// TIA Portal project "PolyMix_v0.1" (V14) (continued)
VERSION : 0.1
   VAR
      DD_Status : Int;
      DD_Mode : Int;
      DD_Alarm : Word;
      DL_Status : Int;
      DL_Mode : Int;
      DL_Alarm : Word;
      Mix_1_Status : Int;
      Mix_1_Mode : Int;
      Mix_1_Alarm : Word;
      Mix_2_Status : Int;
      Mix_2_Mode : Int;
      Mix_2_Alarm : Word;
      Mix_3_Status : Int;
      Mix_3_Mode : Int;
      Mix_3_Alarm : Word;
      KC1_Status : Int;
      Flowmeter : Real;
      Flow_Alarm : Word;
      Level : Real;
      Level_Alarm : Word;
      SP : Real;
      Start : Bool;
      Hand : Bool;
      Warning : Bool;
      Config : Struct
         Use_DD : Bool;   // Использовать сухой дозатор
         Use_DL : Bool;   // Использовать жидкий дозатор
         Use_Mix_1 : Bool;   // Использовать мешалку 1
         Use_Mix_2 : Bool;   // Использовать мешалку 2
         Use_Mix_3 : Bool;   // Использовать мешалку 3
      END_STRUCT;
      Alarm : Word;
   END_VAR
BEGIN
END_DATA_BLOCK

DATA_BLOCK "Time"   // DB13
{ S7_Optimized_Access := 'FALSE' }
VERSION : 0.1
   VAR
      Today : DTL;
      Today_status : Int;
      Set_DTL : DTL;
      Set_status : Int;
      Year : UInt;
      Month : UInt;
      Day : UInt;
      Hour : UInt;
      Minutes : UInt;
      Save : Bool;   // Сохранить время
   END_VAR
BEGIN
END_DATA_BLOCK

// folder: Modules

DATA_BLOCK "DIx_DB"   // DB200
{ S7_Optimized_Access := 'FALSE' }
VERSION : 0.1
// stored: InstanceOfName DIx
"DIx"
BEGIN
END_DATA_BLOCK

DATA_BLOCK "DOx_DB"   // DB201
{ S7_Optimized_Access := 'FALSE' }
VERSION : 0.1
// stored: InstanceOfName DOx
"DOx"
BEGIN
END_DATA_BLOCK

// folder: System blocks/Program resources

DATA_BLOCK "T_Reset"   // DB7
{ S7_Optimized_Access := 'TRUE' }
AUTHOR : Simatic
FAMILY : IEC
NAME : IEC_TMR
VERSION : 1.0
// stored: InstanceOfName IEC_TIMER
"IEC_TIMER"
BEGIN
END_DATA_BLOCK

DATA_BLOCK "clock_5s_ON"   // DB507
{ S7_Optimized_Access := 'TRUE' }
AUTHOR : Simatic
FAMILY : IEC
NAME : IEC_TMR
VERSION : 1.0
// stored: InstanceOfName IEC_TIMER
"IEC_TIMER"
BEGIN
END_DATA_BLOCK

DATA_BLOCK "clock_5s_OFF"   // DB508
{ S7_Optimized_Access := 'TRUE' }
AUTHOR : Simatic
FAMILY : IEC
NAME : IEC_TMR
VERSION : 1.0
// stored: InstanceOfName IEC_TIMER
"IEC_TIMER"
BEGIN
END_DATA_BLOCK

// folder: (top level)

ORGANIZATION_BLOCK "Main"   // OB1, LAD, ProgramCycle
TITLE = "Main Program Sweep (Cycle)"
{ S7_Optimized_Access := 'TRUE' }
VERSION : 0.1
   VAR_INPUT
      Initial_Call : Bool;   // Initial call of this OB
      Remanence : Bool;   // =True, if remanent data are available
   END_VAR
   VAR_TEMP   // added for the SCL form of the ladder/FBD networks
      _w1 : Bool;
   END_VAR
BEGIN

REGION Network 1
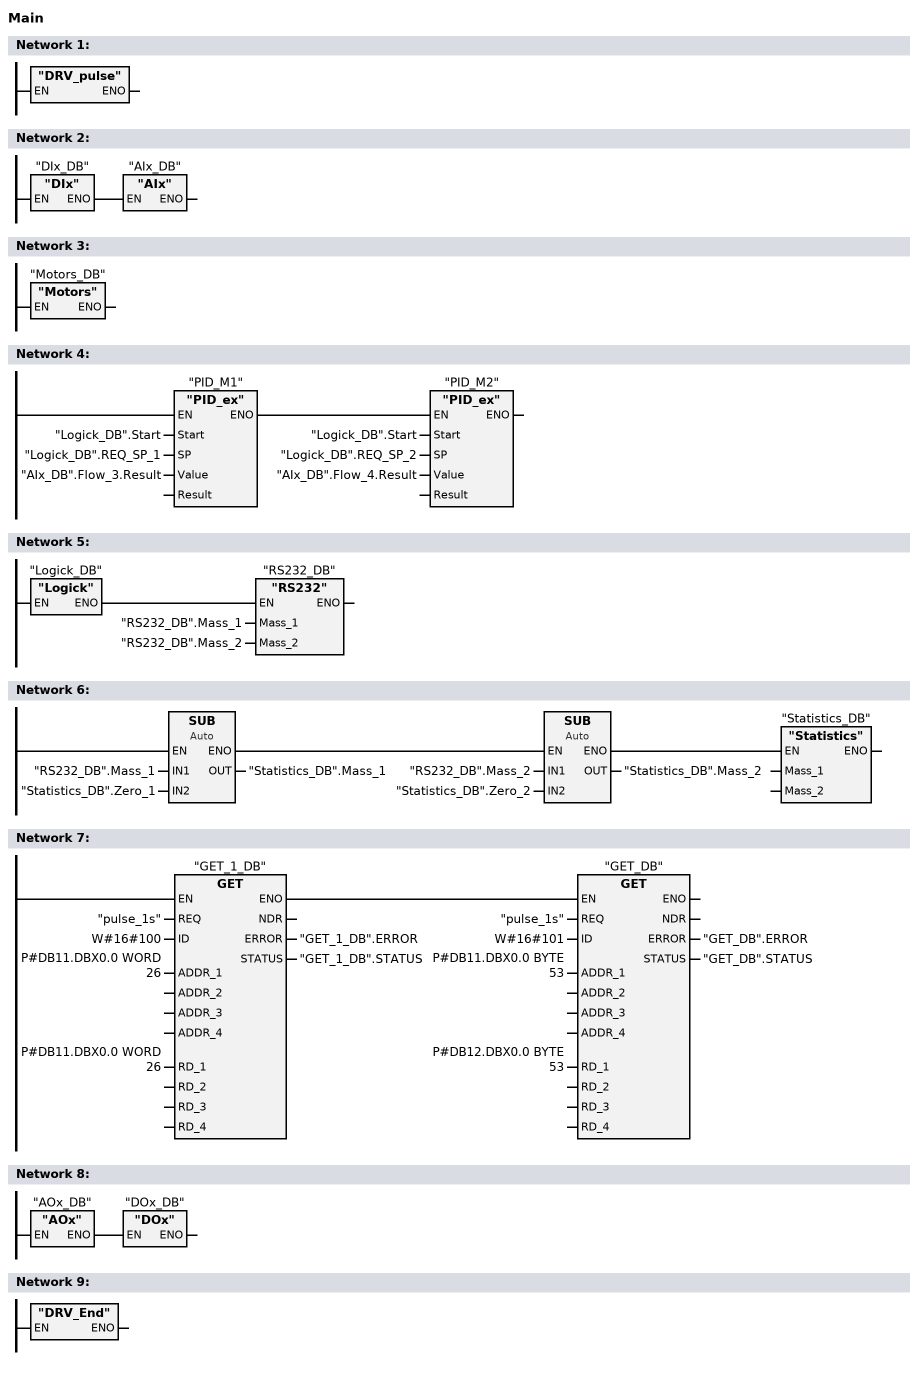
   RUNG wire#powerrail
      "DRV_pulse"()
   END_RUNG
   // the same network as SCL:
   "DRV_pulse"();
END_REGION

REGION Network 2
   RUNG wire#powerrail
      "DIx_DB"()
      "AIx_DB"()
   END_RUNG
   // the same network as SCL:
   "DIx_DB"(ENO => #_w1);   // "DIx"
   IF #_w1 THEN
       "AIx_DB"();   // "AIx"
   END_IF;
END_REGION

REGION Network 3
   RUNG wire#powerrail
      "Motors_DB"()
   END_RUNG
   // the same network as SCL:
   "Motors_DB"();   // "Motors"
END_REGION

REGION Network 4
   RUNG wire#powerrail
      "PID_M1"(Start := "Logick_DB".Start, SP := "Logick_DB".REQ_SP_1, Value := "AIx_DB".Flow_3.Result, Result :=)
      "PID_M2"(Start := "Logick_DB".Start, SP := "Logick_DB".REQ_SP_2, Value := "AIx_DB".Flow_4.Result, Result :=)
   END_RUNG
   // the same network as SCL:
   "PID_M1"(Start := "Logick_DB".Start,   // "PID_ex"
            SP := "Logick_DB".REQ_SP_1,
            Value := "AIx_DB".Flow_3.Result,
            ENO => #_w1);
   IF #_w1 THEN
       "PID_M2"(Start := "Logick_DB".Start, SP := "Logick_DB".REQ_SP_2, Value := "AIx_DB".Flow_4.Result);   // "PID_ex"
   END_IF;
END_REGION

REGION Network 5
   RUNG wire#powerrail
      "Logick_DB"()
      "RS232_DB"(Mass_1 := "RS232_DB".Mass_1, Mass_2 := "RS232_DB".Mass_2)
   END_RUNG
   // the same network as SCL:
   "Logick_DB"(ENO => #_w1);   // "Logick"
   IF #_w1 THEN
       "RS232_DB"(Mass_1 := "RS232_DB".Mass_1, Mass_2 := "RS232_DB".Mass_2);   // "RS232"
   END_IF;
END_REGION

REGION Network 6
   RUNG wire#powerrail
      Sub(in1 := "RS232_DB".Mass_1, in2 := "Statistics_DB".Zero_1, out => "Statistics_DB".Mass_1)
      Sub(in1 := "RS232_DB".Mass_2, in2 := "Statistics_DB".Zero_2, out => "Statistics_DB".Mass_2)
      "Statistics_DB"(Mass_1 :=, Mass_2 :=)
   END_RUNG
   // the same network as SCL:
   "Statistics_DB".Mass_1 := "RS232_DB".Mass_1 - "Statistics_DB".Zero_1;
   "Statistics_DB".Mass_2 := "RS232_DB".Mass_2 - "Statistics_DB".Zero_2;
   "Statistics_DB"();   // "Statistics"
END_REGION

REGION Network 7
   // ENO of a box is taken as its EN; it also drops when the box reports an error
   "GET_1_DB"(REQ := "pulse_1s",   // GET
              ID := W#16#100,
              ADDR_1 := P#DB11.DBX0.0 WORD 26,
              RD_1 := P#DB11.DBX0.0 WORD 26,
              ERROR => "GET_1_DB".ERROR,
              STATUS => "GET_1_DB".STATUS);
   "GET_DB"(REQ := "pulse_1s",   // GET
            ID := W#16#101,
            ADDR_1 := P#DB11.DBX0.0 BYTE 53,
            RD_1 := P#DB12.DBX0.0 BYTE 53,
            ERROR => "GET_DB".ERROR,
            STATUS => "GET_DB".STATUS);
END_REGION

REGION Network 8
   RUNG wire#powerrail
      "AOx_DB"()
      "DOx_DB"()
   END_RUNG
   // the same network as SCL:
   "AOx_DB"(ENO => #_w1);   // "AOx"
   IF #_w1 THEN
       "DOx_DB"();   // "DOx"
   END_IF;
END_REGION

REGION Network 9
   RUNG wire#powerrail
      "DRV_End"()
   END_RUNG
   // the same network as SCL:
   "DRV_End"();
END_REGION
END_ORGANIZATION_BLOCK

ORGANIZATION_BLOCK "Time error interrupt"   // OB80, LAD, TimeErrorInterrupt
{ S7_Optimized_Access := 'TRUE' }
VERSION : 0.1
   VAR_INPUT
      Fault_ID : Byte;   // Fault identifier
      Csg_OBnr : OB_Any;   // Number of OB causing the error
      Csg_Prio : UInt;   // Priority of OB causing the error
   END_VAR
BEGIN
END_ORGANIZATION_BLOCK

ORGANIZATION_BLOCK "Diagnostic error interrupt"   // OB82, LAD, DiagnosticErrorInterrupt
{ S7_Optimized_Access := 'TRUE' }
VERSION : 0.1
   VAR_INPUT
      IO_State : Word;   // IO state of the HW object
      LADDR : Hw_Any;   // Hardware identifier
      Channel : UInt;   // Channel number
      MultiError : Bool;   // =true if more than one error is present
   END_VAR
BEGIN
END_ORGANIZATION_BLOCK

ORGANIZATION_BLOCK "Startup"   // OB100, LAD, Startup
TITLE = "Complete Restart"
{ S7_Optimized_Access := 'TRUE' }
VERSION : 0.1
   VAR_INPUT
      LostRetentive : Bool;   // True if retentive data are lost
      LostRTC : Bool;   // True if date and time are lost
   END_VAR
BEGIN

REGION Network 1: Запуск автоматики
END_REGION

REGION Network 2
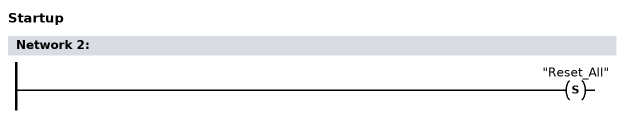
   RUNG wire#powerrail
      S_Coil( "Reset_All" )
   END_RUNG
   // the same network as SCL:
   "Reset_All" := TRUE;
END_REGION
END_ORGANIZATION_BLOCK

// folder: DRV_Low

FUNCTION_BLOCK "DI_ex"   // FB100, LAD
{ S7_Optimized_Access := 'FALSE' }
VERSION : 0.1
   VAR_INPUT
      Input : Bool;   // Входящий сигнал
      pulse : Bool;   // Частота фильтрации дребезка
   END_VAR
   VAR_OUTPUT
      Signal : Bool;   // Результирующий сигнал
   END_VAR
   VAR
      Hand : Bool;   // 0 - Авто, 1 - Ручной
      Start_M : Bool;   // Запуск в ручном режиме
      Data : Bool;   // Отфильтрованный сигнал
      Inverse : Bool;   // Инверсия входного сигнала
      Filter_On : Struct   // Фильтр наличия сигнала
         SP : Int;
         Now : Int;
         "Exit" : Bool;
         Start : Bool;
         Pause : Bool;
         Reset : Bool;
      END_STRUCT;
      Filter_Off : Struct   // Фильтр отсутствия сигнала
         SP : Int;
         Now : Int;
         "Exit" : Bool;
         Start : Bool;
         Pause : Bool;
         Reset : Bool;
      END_STRUCT;
      res_1 : Word;
   END_VAR
   VAR_TEMP   // added for the SCL form of the ladder/FBD networks
      _w1 : Bool;
   END_VAR
BEGIN

REGION Network 1: Устройство в ручном режиме
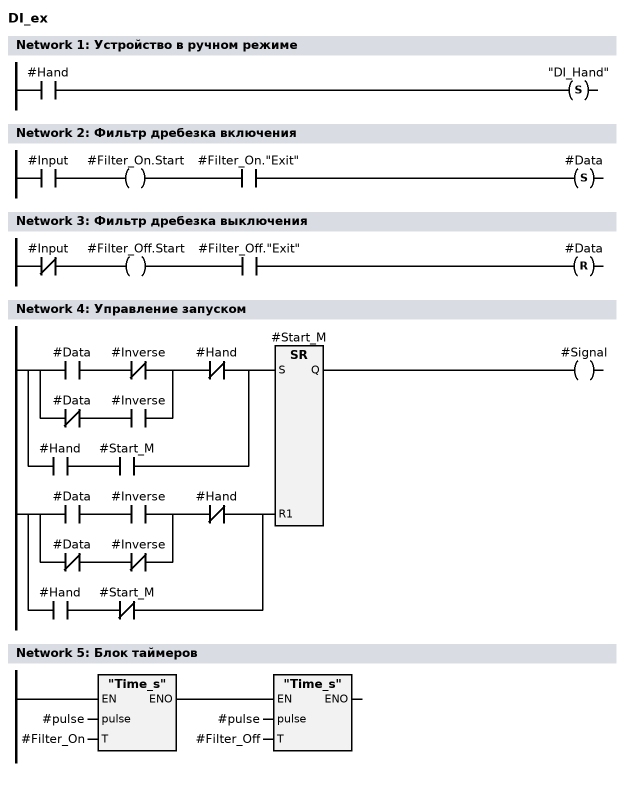
   RUNG wire#powerrail
      Contact( #Hand )
      S_Coil( "DI_Hand" )
   END_RUNG
   // the same network as SCL:
   IF #Hand THEN "DI_Hand" := TRUE; END_IF;
END_REGION

REGION Network 2: Фильтр дребезка включения
   RUNG wire#powerrail
      Contact( #Input )
      Coil( #Filter_On.Start )
      Contact( #Filter_On."Exit" )
      S_Coil( #Data )
   END_RUNG
   // the same network as SCL:
   #Filter_On.Start := #Input;
   IF #Input AND #Filter_On."Exit" THEN #Data := TRUE; END_IF;
END_REGION

REGION Network 3: Фильтр дребезка выключения
   RUNG wire#powerrail
      I_Contact( #Input )
      Coil( #Filter_Off.Start )
      Contact( #Filter_Off."Exit" )
      R_Coil( #Data )
   END_RUNG
   // the same network as SCL:
   #Filter_Off.Start := NOT #Input;
   IF NOT #Input AND #Filter_Off."Exit" THEN #Data := FALSE; END_IF;
END_REGION

REGION Network 4: Управление запуском
   RUNG wire#powerrail
      Contact( #Data )
      I_Contact( #Inverse )
      wire#w1
      I_Contact( #Hand )
      wire#w2
      S_SR(operand := #Start_M, r1 := wire#w4)
      Coil( #Signal )
   END_RUNG
   RUNG wire#powerrail
      I_Contact( #Data )
      Contact( #Inverse )
   END_RUNG wire#w1
   RUNG wire#powerrail
      Contact( #Hand )
      Contact( #Start_M )
   END_RUNG wire#w2
   RUNG wire#powerrail
      Contact( #Data )
      Contact( #Inverse )
      wire#w3
      I_Contact( #Hand )
   END_RUNG wire#w4
   RUNG wire#powerrail
      I_Contact( #Data )
      I_Contact( #Inverse )
   END_RUNG wire#w3
   RUNG wire#powerrail
      Contact( #Hand )
      I_Contact( #Start_M )
   END_RUNG wire#w4
   // the same network as SCL:
   #_w1 := (((#Data AND #Inverse) OR (NOT #Data AND NOT #Inverse)) AND NOT #Hand) OR (#Hand AND NOT #Start_M);
   IF (((#Data AND NOT #Inverse) OR (NOT #Data AND #Inverse)) AND NOT #Hand) OR (#Hand AND #Start_M) THEN
       #Start_M := TRUE;   // SR flip-flop
   END_IF;
   IF #_w1 THEN #Start_M := FALSE; END_IF;
   #Signal := #Start_M;
END_REGION

REGION Network 5: Блок таймеров
   RUNG wire#powerrail
      "Time_s"(pulse := #pulse, T := #Filter_On)
      "Time_s"(pulse := #pulse, T := #Filter_Off)
   END_RUNG
   // the same network as SCL:
   "Time_s"(pulse := #pulse, T := #Filter_On, ENO => #_w1);
   IF #_w1 THEN "Time_s"(pulse := #pulse, T := #Filter_Off); END_IF;
END_REGION
END_FUNCTION_BLOCK

FUNCTION_BLOCK "DO_ex"   // FB101, LAD
{ S7_Optimized_Access := 'FALSE' }
VERSION : 0.1
   VAR_IN_OUT
      Start_A : Bool;   // Управляющий сигнал из программы
      pulse : Bool;   // Частота длительности импульса
      Q : Bool;   // Выходной сигнал контроллера
   END_VAR
   VAR
      Hand : Bool;   // 0 - Авто, 1 - Ручной
      Start_M : Bool;   // Запуск в ручном режиме
      Simulation : Bool;   // Режим симуляции
      Inverse : Bool;   // Инверсия выхода
      Impulse : Bool;   // Импульсный режим
      T_Impulse : Struct   // Длительность импульса
         SP : Int := 5;
         Now : Int;
         "Exit" : Bool;
         Start : Bool;
         Pause : Bool;
         Reset : Bool;
      END_STRUCT;
   END_VAR
   VAR_TEMP   // added for the SCL form of the ladder/FBD networks
      _w1 : Bool;
   END_VAR
BEGIN

REGION Network 1: Устройство в ручном режиме
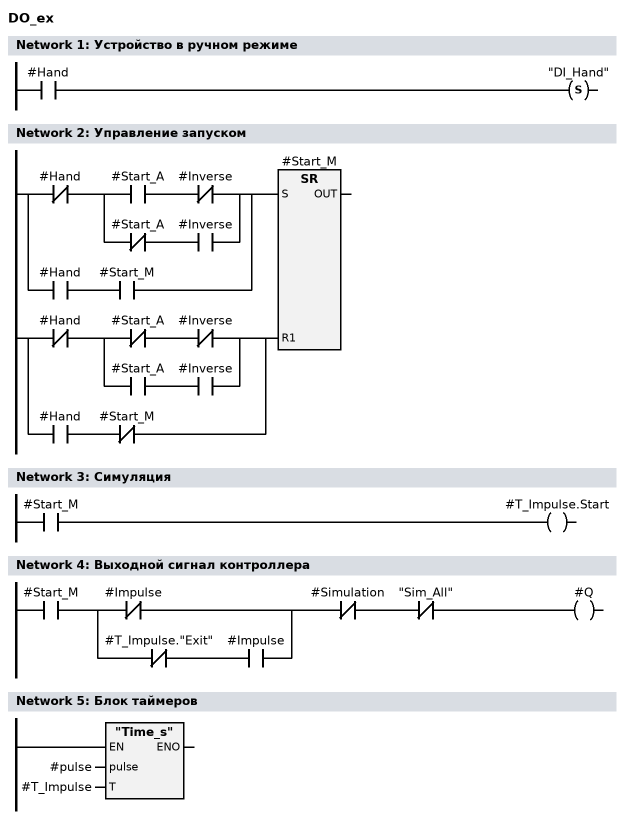
   RUNG wire#powerrail
      Contact( #Hand )
      S_Coil( "DI_Hand" )
   END_RUNG
   // the same network as SCL:
   IF #Hand THEN "DI_Hand" := TRUE; END_IF;
END_REGION

REGION Network 2: Управление запуском
   RUNG wire#powerrail
      I_Contact( #Hand )
      wire#w1
      Contact( #Start_A )
      I_Contact( #Inverse )
      wire#w2
      S_SR(operand := #Start_M, r1 := wire#w4)
   END_RUNG
   RUNG wire#w1
      I_Contact( #Start_A )
      Contact( #Inverse )
   END_RUNG wire#w2
   RUNG wire#powerrail
      Contact( #Hand )
      Contact( #Start_M )
   END_RUNG wire#w2
   RUNG wire#powerrail
      I_Contact( #Hand )
      wire#w3
      I_Contact( #Start_A )
      I_Contact( #Inverse )
   END_RUNG wire#w4
   RUNG wire#w3
      Contact( #Start_A )
      Contact( #Inverse )
   END_RUNG wire#w4
   RUNG wire#powerrail
      Contact( #Hand )
      I_Contact( #Start_M )
   END_RUNG wire#w4
   // the same network as SCL:
   #_w1 := (NOT #Hand AND ((NOT #Start_A AND NOT #Inverse) OR (#Start_A AND #Inverse))) OR (#Hand AND NOT #Start_M);
   IF (NOT #Hand AND ((#Start_A AND NOT #Inverse) OR (NOT #Start_A AND #Inverse))) OR (#Hand AND #Start_M) THEN
       #Start_M := TRUE;   // SR flip-flop
   END_IF;
   IF #_w1 THEN #Start_M := FALSE; END_IF;
END_REGION

REGION Network 3: Симуляция
   RUNG wire#powerrail
      Contact( #Start_M )
      Coil( #T_Impulse.Start )
   END_RUNG
   // the same network as SCL:
   #T_Impulse.Start := #Start_M;
END_REGION

REGION Network 4: Выходной сигнал контроллера
   RUNG wire#powerrail
      Contact( #Start_M )
      wire#w1
      I_Contact( #Impulse )
      wire#w2
      I_Contact( #Simulation )
      I_Contact( "Sim_All" )
      Coil( #Q )
   END_RUNG
   RUNG wire#w1
      I_Contact( #T_Impulse."Exit" )
      Contact( #Impulse )
   END_RUNG wire#w2
   // the same network as SCL:
   #Q := #Start_M AND (NOT #Impulse OR (NOT #T_Impulse."Exit" AND #Impulse)) AND NOT #Simulation AND NOT "Sim_All";
END_REGION

REGION Network 5: Блок таймеров
   RUNG wire#powerrail
      "Time_s"(pulse := #pulse, T := #T_Impulse)
   END_RUNG
   // the same network as SCL:
   "Time_s"(pulse := #pulse, T := #T_Impulse);
END_REGION
END_FUNCTION_BLOCK

FUNCTION_BLOCK "DRV_Micro"   // FB104, LAD
{ S7_Optimized_Access := 'FALSE' }
VERSION : 0.1
   VAR_INPUT
      Start_A : Bool;   // Запрос запуска
      FB : Bool;   // ОС
      Reset : Bool;   // Сброс аварий
      All_Block : Bool;   // Блокировка
   END_VAR
   VAR_OUTPUT
      CMD : Bool;   // Команда
   END_VAR
   VAR_IN_OUT
      Alarm : Bool;   // Авария
   END_VAR
   VAR
      Hand : Bool;   // Ручной режим
      Start_M : Bool;   // Запуск в ручном режиме
      No_FB : Bool;   // Не использовать ОС
      ON : Bool;   // Успешно запущено
      OFF : Bool;   // Успешно остановлено
      Status : Int;   // Статус устройства / Статус привода
      Wait_On : Struct   // Ожидание ОС контактора / Время на запуск
         SP : Int := 2;
         Now : Int;
         "Exit" : Bool;
         Start : Bool;
         Pause : Bool;
         Reset : Bool;
      END_STRUCT;
      Wait_Off : Struct   // Ожидание концевиков / Время на останов
         SP : Int := 2;
         Now : Int;
         "Exit" : Bool;
         Start : Bool;
         Pause : Bool;
         Reset : Bool;
      END_STRUCT;
   END_VAR
   VAR_TEMP   // added for the SCL form of the ladder/FBD networks
      _w1 : Bool;
      _w2 : Bool;
   END_VAR
BEGIN

REGION Network 1: Управление запуском / дискретный управляющий сигнал
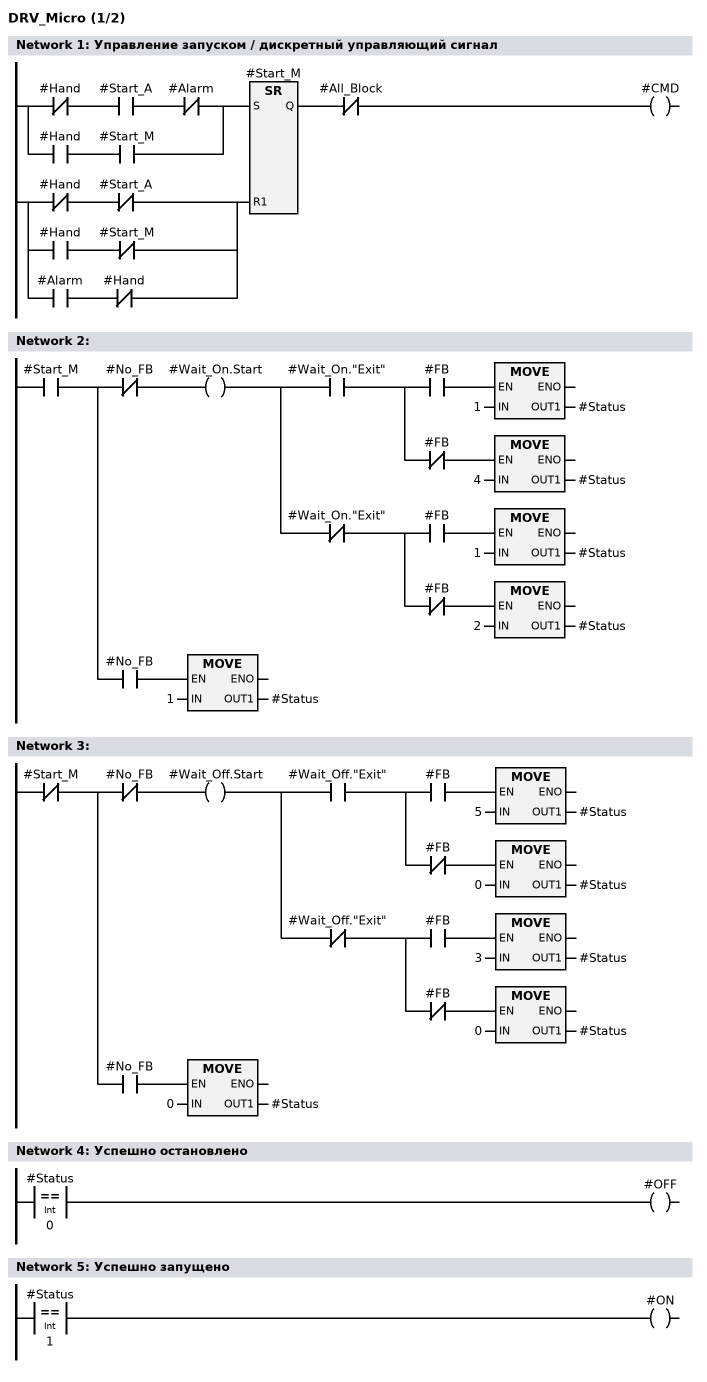
   RUNG wire#powerrail
      I_Contact( #Hand )
      Contact( #Start_A )
      I_Contact( #Alarm )
      wire#w1
      S_SR(operand := #Start_M, r1 := wire#w2)
      I_Contact( #All_Block )
      Coil( #CMD )
   END_RUNG
   RUNG wire#powerrail
      Contact( #Hand )
      Contact( #Start_M )
   END_RUNG wire#w1
   RUNG wire#powerrail
      I_Contact( #Hand )
      I_Contact( #Start_A )
   END_RUNG wire#w2
   RUNG wire#powerrail
      Contact( #Hand )
      I_Contact( #Start_M )
   END_RUNG wire#w2
   RUNG wire#powerrail
      Contact( #Alarm )
      I_Contact( #Hand )
   END_RUNG wire#w2
   // the same network as SCL:
   #_w1 := (NOT #Hand AND NOT #Start_A) OR (#Hand AND NOT #Start_M) OR (#Alarm AND NOT #Hand);
   IF (NOT #Hand AND #Start_A AND NOT #Alarm) OR (#Hand AND #Start_M) THEN
       #Start_M := TRUE;   // SR flip-flop
   END_IF;
   IF #_w1 THEN #Start_M := FALSE; END_IF;
   #CMD := #Start_M AND NOT #All_Block;
END_REGION

REGION Network 2
   RUNG wire#powerrail
      Contact( #Start_M )
      wire#w1
      I_Contact( #No_FB )
      Coil( #Wait_On.Start )
      wire#w2
      Contact( #Wait_On."Exit" )
      wire#w3
      Contact( #FB )
      Move(in := 1, out1 => #Status)
   END_RUNG
   RUNG wire#w3
      I_Contact( #FB )
      Move(in := 4, out1 => #Status)
   END_RUNG
   RUNG wire#w2
      I_Contact( #Wait_On."Exit" )
      wire#w4
      Contact( #FB )
      Move(in := 1, out1 => #Status)
   END_RUNG
   RUNG wire#w4
      I_Contact( #FB )
      Move(in := 2, out1 => #Status)
   END_RUNG
   RUNG wire#w1
      Contact( #No_FB )
      Move(in := 1, out1 => #Status)
   END_RUNG
   // the same network as SCL:
   #Wait_On.Start := #Start_M AND NOT #No_FB;
   #_w1 := #Wait_On.Start AND #Wait_On."Exit";
   IF #_w1 AND #FB THEN #Status := 1; END_IF;
   IF #_w1 AND NOT #FB THEN #Status := 4; END_IF;
   #_w2 := #Wait_On.Start AND NOT #Wait_On."Exit";
   IF #_w2 AND #FB THEN #Status := 1; END_IF;
   IF #_w2 AND NOT #FB THEN #Status := 2; END_IF;
   IF #Start_M AND #No_FB THEN #Status := 1; END_IF;
END_REGION

REGION Network 3
   RUNG wire#powerrail
      I_Contact( #Start_M )
      wire#w1
      I_Contact( #No_FB )
      Coil( #Wait_Off.Start )
      wire#w2
      Contact( #Wait_Off."Exit" )
      wire#w3
      Contact( #FB )
      Move(in := 5, out1 => #Status)
   END_RUNG
   RUNG wire#w3
      I_Contact( #FB )
      Move(in := 0, out1 => #Status)
   END_RUNG
   RUNG wire#w2
      I_Contact( #Wait_Off."Exit" )
      wire#w4
      Contact( #FB )
      Move(in := 3, out1 => #Status)
   END_RUNG
   RUNG wire#w4
      I_Contact( #FB )
      Move(in := 0, out1 => #Status)
   END_RUNG
   RUNG wire#w1
      Contact( #No_FB )
      Move(in := 0, out1 => #Status)
   END_RUNG
   // the same network as SCL:
   #Wait_Off.Start := NOT #Start_M AND NOT #No_FB;
   #_w1 := #Wait_Off.Start AND #Wait_Off."Exit";
   IF #_w1 AND #FB THEN #Status := 5; END_IF;
   IF #_w1 AND NOT #FB THEN #Status := 0; END_IF;
   #_w2 := #Wait_Off.Start AND NOT #Wait_Off."Exit";
   IF #_w2 AND #FB THEN #Status := 3; END_IF;
   IF #_w2 AND NOT #FB THEN #Status := 0; END_IF;
   IF NOT #Start_M AND #No_FB THEN #Status := 0; END_IF;
END_REGION

REGION Network 4: Успешно остановлено
   RUNG wire#powerrail
      { S7_Templates := "SrcType := Int" } EQ_Contact(in1 := #Status, in2 := 0)
      Coil( #OFF )
   END_RUNG
   // the same network as SCL:
   #OFF := #Status = 0;
END_REGION

REGION Network 5: Успешно запущено
   RUNG wire#powerrail
      { S7_Templates := "SrcType := Int" } EQ_Contact(in1 := #Status, in2 := 1)
      Coil( #ON )
   END_RUNG
   // the same network as SCL:
   #ON := #Status = 1;
END_REGION

REGION Network 6: Авария
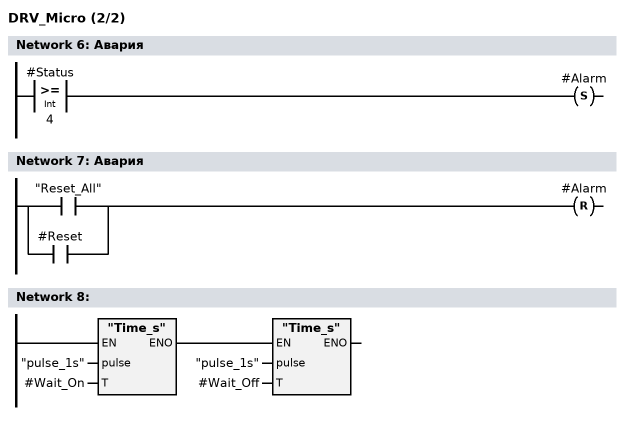
   RUNG wire#powerrail
      { S7_Templates := "SrcType := Int" } GE_Contact(in1 := #Status, in2 := 4)
      S_Coil( #Alarm )
   END_RUNG
   // the same network as SCL:
   IF #Status >= 4 THEN #Alarm := TRUE; END_IF;
END_REGION

REGION Network 7: Авария
   RUNG wire#powerrail
      Contact( "Reset_All" )
      wire#w1
      R_Coil( #Alarm )
   END_RUNG
   RUNG wire#powerrail
      Contact( #Reset )
   END_RUNG wire#w1
   // the same network as SCL:
   IF "Reset_All" OR #Reset THEN #Alarm := FALSE; END_IF;
END_REGION

REGION Network 8
   RUNG wire#powerrail
      "Time_s"(pulse := "pulse_1s", T := #Wait_On)
      "Time_s"(pulse := "pulse_1s", T := #Wait_Off)
   END_RUNG
   // the same network as SCL:
   "Time_s"(pulse := "pulse_1s", T := #Wait_On, ENO => #_w1);
   IF #_w1 THEN "Time_s"(pulse := "pulse_1s", T := #Wait_Off); END_IF;
END_REGION
END_FUNCTION_BLOCK

// folder: Modules

FUNCTION_BLOCK "DIx"   // FB200, LAD
{ S7_Optimized_Access := 'FALSE' }
VERSION : 0.1
// Input - входной сигнал контроллера
// pulse - частота фильтрации дребезга
// Signal - обработанный и отфильтрованный сигнал, используемый в дальнейшем
   VAR
      M1_QF : "DI_ex";
      M2_QF : "DI_ex";
      M3_QF : "DI_ex";
      Heat_1 : "DI_ex";
      Heat_2 : "DI_ex";
      Heat_3 : "DI_ex";
      Heat_4 : "DI_ex";
      AllBlock : "DI_ex";
      Mass_1 : "DI_ex";
      Mass_2 : "DI_ex";
   END_VAR
   VAR_TEMP   // added for the SCL form of the ladder/FBD networks
      _w1 : Bool;
      _w2 : Bool;
      _w3 : Bool;
   END_VAR
BEGIN

REGION Network 1
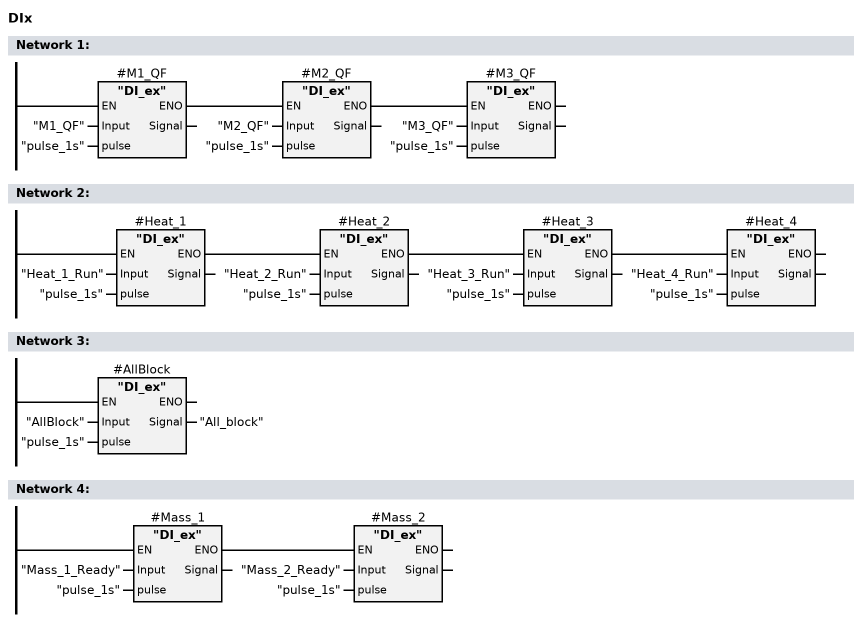
   RUNG wire#powerrail
      #M1_QF(Input := "M1_QF", pulse := "pulse_1s", Signal =>)
      #M2_QF(Input := "M2_QF", pulse := "pulse_1s", Signal =>)
      #M3_QF(Input := "M3_QF", pulse := "pulse_1s", Signal =>)
   END_RUNG
   // the same network as SCL:
   #M1_QF(Input := "M1_QF", pulse := "pulse_1s", ENO => #_w1);   // "DI_ex"
   #M2_QF(EN := #_w1, Input := "M2_QF", pulse := "pulse_1s", ENO => #_w2);   // "DI_ex"
   IF #_w2 THEN
       #M3_QF(Input := "M3_QF", pulse := "pulse_1s");   // "DI_ex"
   END_IF;
END_REGION

REGION Network 2
   RUNG wire#powerrail
      #Heat_1(Input := "Heat_1_Run", pulse := "pulse_1s", Signal =>)
      #Heat_2(Input := "Heat_2_Run", pulse := "pulse_1s", Signal =>)
      #Heat_3(Input := "Heat_3_Run", pulse := "pulse_1s", Signal =>)
      #Heat_4(Input := "Heat_4_Run", pulse := "pulse_1s", Signal =>)
   END_RUNG
   // the same network as SCL:
   #Heat_1(Input := "Heat_1_Run", pulse := "pulse_1s", ENO => #_w1);   // "DI_ex"
   #Heat_2(EN := #_w1, Input := "Heat_2_Run", pulse := "pulse_1s", ENO => #_w2);   // "DI_ex"
   #Heat_3(EN := #_w2, Input := "Heat_3_Run", pulse := "pulse_1s", ENO => #_w3);   // "DI_ex"
   IF #_w3 THEN
       #Heat_4(Input := "Heat_4_Run", pulse := "pulse_1s");   // "DI_ex"
   END_IF;
END_REGION

REGION Network 3
   RUNG wire#powerrail
      #AllBlock(Input := "AllBlock", pulse := "pulse_1s", Signal => "All_block")
   END_RUNG
   // the same network as SCL:
   #AllBlock(Input := "AllBlock", pulse := "pulse_1s", Signal => "All_block");   // "DI_ex"
END_REGION

REGION Network 4
   RUNG wire#powerrail
      #Mass_1(Input := "Mass_1_Ready", pulse := "pulse_1s", Signal =>)
      #Mass_2(Input := "Mass_2_Ready", pulse := "pulse_1s", Signal =>)
   END_RUNG
   // the same network as SCL:
   #Mass_1(Input := "Mass_1_Ready", pulse := "pulse_1s", ENO => #_w1);   // "DI_ex"
   IF #_w1 THEN
       #Mass_2(Input := "Mass_2_Ready", pulse := "pulse_1s");   // "DI_ex"
   END_IF;
END_REGION
END_FUNCTION_BLOCK

FUNCTION_BLOCK "DOx"   // FB201, LAD
{ S7_Optimized_Access := 'FALSE' }
VERSION : 0.1
// Start - управляющий сигнал из программы
// Q - выходной сигнал контроллера
// pulse - кратность времени в импульсном режиме
   VAR
      M1_CMD : "DO_ex";
      M2_CMD : "DO_ex";
      M3_CMD : "DO_ex";
      LED_Error_1 : "DO_ex";
      LED_Error_2 : "DO_ex";
      LED_Alarm : "DO_ex";
      LED_M1_Alarm : "DO_ex";
      LED_M2_Alarm : "DO_ex";
      LED_M3_Alarm : "DO_ex";
   END_VAR
   VAR_TEMP   // added for the SCL form of the ladder/FBD networks
      _w1 : Bool;
      _w2 : Bool;
   END_VAR
BEGIN

REGION Network 1: Насосы
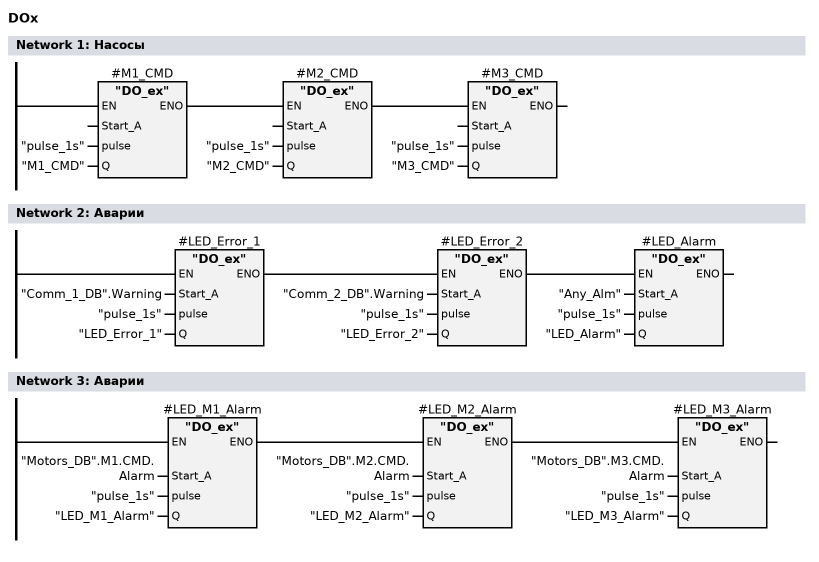
   RUNG wire#powerrail
      #M1_CMD(Start_A :=, pulse := "pulse_1s", Q := "M1_CMD")
      #M2_CMD(Start_A :=, pulse := "pulse_1s", Q := "M2_CMD")
      #M3_CMD(Start_A :=, pulse := "pulse_1s", Q := "M3_CMD")
   END_RUNG
   // the same network as SCL:
   #M1_CMD(pulse := "pulse_1s", Q := "M1_CMD", ENO => #_w1);   // "DO_ex"
   #M2_CMD(EN := #_w1, pulse := "pulse_1s", Q := "M2_CMD", ENO => #_w2);   // "DO_ex"
   IF #_w2 THEN
       #M3_CMD(pulse := "pulse_1s", Q := "M3_CMD");   // "DO_ex"
   END_IF;
END_REGION

REGION Network 2: Аварии
   RUNG wire#powerrail
      #LED_Error_1(Start_A := "Comm_1_DB".Warning, pulse := "pulse_1s", Q := "LED_Error_1")
      #LED_Error_2(Start_A := "Comm_2_DB".Warning, pulse := "pulse_1s", Q := "LED_Error_2")
      #LED_Alarm(Start_A := "Any_Alm", pulse := "pulse_1s", Q := "LED_Alarm")
   END_RUNG
   // the same network as SCL:
   #LED_Error_1(Start_A := "Comm_1_DB".Warning, pulse := "pulse_1s", Q := "LED_Error_1", ENO => #_w1);   // "DO_ex"
   #LED_Error_2(EN := #_w1,   // "DO_ex"
                Start_A := "Comm_2_DB".Warning,
                pulse := "pulse_1s",
                Q := "LED_Error_2",
                ENO => #_w2);
   IF #_w2 THEN
       #LED_Alarm(Start_A := "Any_Alm", pulse := "pulse_1s", Q := "LED_Alarm");   // "DO_ex"
   END_IF;
END_REGION

REGION Network 3: Аварии
   RUNG wire#powerrail
      #LED_M1_Alarm(Start_A := "Motors_DB".M1.CMD.Alarm, pulse := "pulse_1s", Q := "LED_M1_Alarm")
      #LED_M2_Alarm(Start_A := "Motors_DB".M2.CMD.Alarm, pulse := "pulse_1s", Q := "LED_M2_Alarm")
      #LED_M3_Alarm(Start_A := "Motors_DB".M3.CMD.Alarm, pulse := "pulse_1s", Q := "LED_M3_Alarm")
   END_RUNG
   // the same network as SCL:
   #LED_M1_Alarm(Start_A := "Motors_DB".M1.CMD.Alarm, pulse := "pulse_1s", Q := "LED_M1_Alarm", ENO => #_w1);   // "DO_ex"
   #LED_M2_Alarm(EN := #_w1,   // "DO_ex"
                 Start_A := "Motors_DB".M2.CMD.Alarm,
                 pulse := "pulse_1s",
                 Q := "LED_M2_Alarm",
                 ENO => #_w2);
   IF #_w2 THEN
       #LED_M3_Alarm(Start_A := "Motors_DB".M3.CMD.Alarm, pulse := "pulse_1s", Q := "LED_M3_Alarm");   // "DO_ex"
   END_IF;
END_REGION
END_FUNCTION_BLOCK

// folder: System

FUNCTION_BLOCK "PID_ex"   // FB99, LAD
{ S7_Optimized_Access := 'FALSE' }
VERSION : 0.1
   VAR_INPUT
      Start : Bool;   // Команда запуска
      SP : Real;   // Уставка
      Value : Real;   // Показания датчика
   END_VAR
   VAR_IN_OUT
      Result : Real;   // Управляющее воздействие
   END_VAR
   VAR
      Hand : Bool;   // Ручной режим
      Err_Ack : Bool;   // Подтверждение аварии
      Reset : Bool;   // Сброс ПИД
      Error : Bool;   // Авария ПИД
      Invert : Bool;   // Инверсия работы
      SP_H : Bool;   // Авария уставки - превышение
      SP_L : Bool;   // Авария уставки - занижение
      In_H : Bool;   // Авария датчика - превышение
      In_L : Bool;   // Авария датчика - занижение
      Activate : Bool;   // Активировать ПИД
      Error_code : DWord;   // Код аварии
      Warning_code : DWord;   // Код предупреждения
      HandValue : Real;   // Выход ПИД в ручном режиме
      SP_P : Real := 1.5;   // Коэффициент пропорциональности
      SP_Ti : Real := 150.0;   // Время интегрирования
      SP_Td : Real;   // Время дифференцирования
      SP_Cycle : Real := 0.2;   // Время цикла
      Disturvance : Real;   // Внешнее воздействие
      Max_SP : Real := 500.0;   // Максимальное значение уставки
      Min_SP : Real := -500.0;   // Минимальное значение уставки
      Max_in : Real := 500.0;   // Максимальное значение датчика
      Min_in : Real := -500.0;   // Минимальное значение датчика
      Max_out : Real := 100.0;   // Максимальное значение выхода
      Min_out : Real := 0.0;   // Минимальное значение выхода
      "Type" : Int := 1;   // Режим работы
      State : Int;   // Состояние
      Mode : Int := 3;   // Режим
      PID : PID_Compact;   // ПИД
      DeadBand : Real;   // Мёртвая зона
      Max : Real;   // Верняя граница мёртвой зоны
      Min : Real;   // Нижняя граница мёртвой зоны
      Converter : Struct
         Use_Min_In : Bool;   // Отсекать входные значения ниже минимума
         Use_Max_In : Bool;   // Отсекать входные значения выше максимума
         Use_Min_Out : Bool;   // Отсекать результат ниже минимума
         Use_Max_Out : Bool;   // Отсекать результат выше максимума
         IO : Bool;   // Входной/Выходной режим
         Inverse : Bool;   // Инверсия выхода
         Min_In : Real := 0.0;   // Минимальный входной сигнал
         Max_In : Real := 100.0;   // Максимальный входной сигнал
         Min_Out : Real;   // Минимальный выходной сигнал
         Max_Out : Real;   // Максимальный выходной сигнал
      END_STRUCT;
      Conveter_Back : Struct
         Use_Min_In : Bool;   // Отсекать входные значения ниже минимума
         Use_Max_In : Bool;   // Отсекать входные значения выше максимума
         Use_Min_Out : Bool;   // Отсекать результат ниже минимума
         Use_Max_Out : Bool;   // Отсекать результат выше максимума
         IO : Bool;   // Входной/Выходной режим
         Inverse : Bool;   // Инверсия выхода
         Min_In : Real;   // Минимальный входной сигнал
         Max_In : Real;   // Максимальный входной сигнал
         Min_Out : Real := 0.0;   // Минимальный выходной сигнал
         Max_Out : Real := 100.0;   // Максимальный выходной сигнал
      END_STRUCT;
      C : Struct
         SP : Real := 1.0;   // Уставка
         Now : Real;   // Текущий счёт
         One : Real;   // Вес импульса
         Progress : Real;   // Прогресс выполнения
         "Exit" : Bool;   // Счёт завершён
         Start : Bool;   // Запуск
         Pause : Bool;   // Пауза
         Reset : Bool;   // Сброс счёта
         pos : Bool;   // Контроль фронта сигнала
      END_STRUCT;
   END_VAR
   VAR_TEMP
      PID_Output : Real;
   END_VAR
   VAR_TEMP   // added for the SCL form of the ladder/FBD networks
      _w1 : Bool;
   END_VAR
BEGIN

REGION Network 1: Сброс ПИД
